// TIA Portal project "liquid refill system" (V18) (continued)
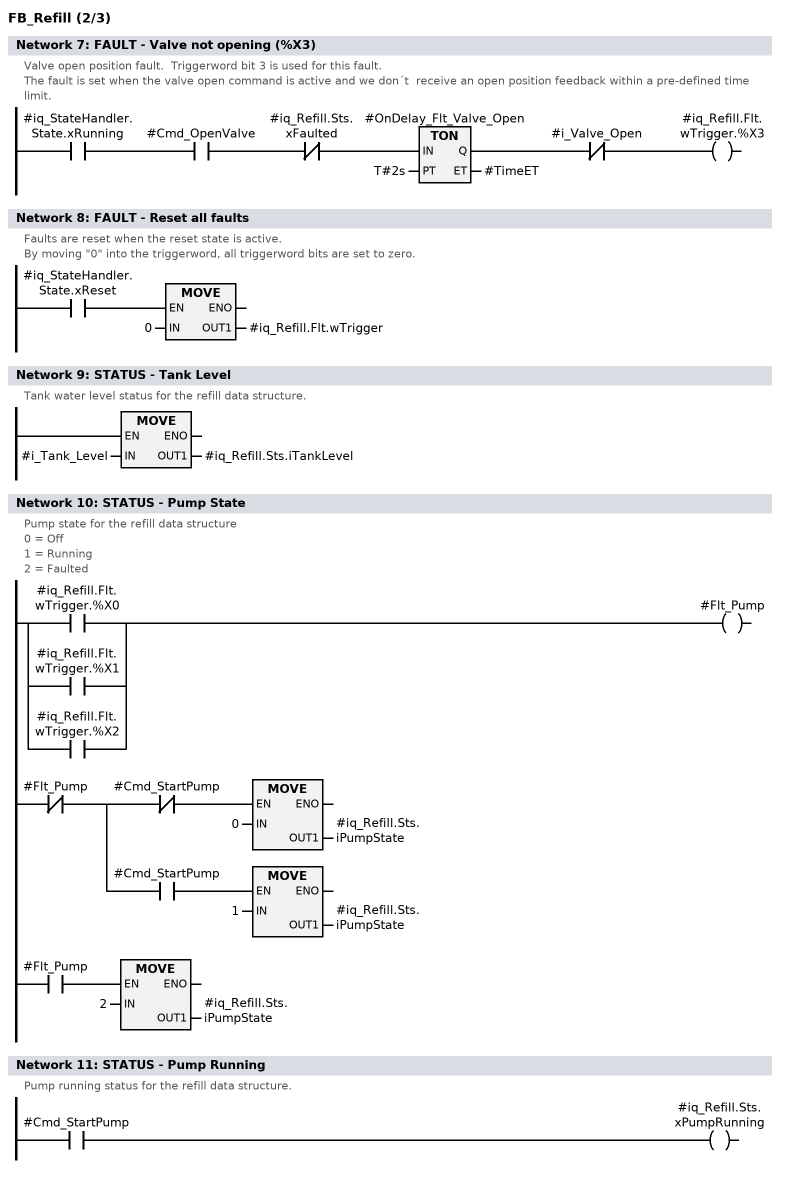
   #OnDelay_Flt_Valve_Open.TON(IN := #iq_StateHandler.State.xRunning AND #Cmd_OpenValve AND NOT #iq_Refill.Sts.xFaulted,
                           PT := T#2s,
                           ET => #TimeET);
   #iq_Refill.Flt.wTrigger.%X3 := #OnDelay_Flt_Valve_Open.Q AND NOT #i_Valve_Open;
END_REGION

REGION Network 8: FAULT - Reset all faults
   // Faults are reset when the reset state is active.
   // By moving "0" into the triggerword, all triggerword bits are set to zero.
   RUNG wire#powerrail
      Contact( #iq_StateHandler.State.xReset )
      Move(in := 0, out1 => #iq_Refill.Flt.wTrigger)
   END_RUNG
   // the same network as SCL:
   IF #iq_StateHandler.State.xReset THEN #iq_Refill.Flt.wTrigger := 0; END_IF;
END_REGION

REGION Network 9: STATUS - Tank Level
   // Tank water level status for the refill data structure.
   RUNG wire#powerrail
      Move(in := #i_Tank_Level, out1 => #iq_Refill.Sts.iTankLevel)
   END_RUNG
   // the same network as SCL:
   #iq_Refill.Sts.iTankLevel := #i_Tank_Level;
END_REGION

REGION Network 10: STATUS - Pump State
   // Pump state for the refill data structure
   // 0 = Off
   // 1 = Running
   // 2 = Faulted
   RUNG wire#powerrail
      Contact( #iq_Refill.Flt.wTrigger.%X0 )
      wire#w1
      Coil( #Flt_Pump )
   END_RUNG
   RUNG wire#powerrail
      Contact( #iq_Refill.Flt.wTrigger.%X1 )
   END_RUNG wire#w1
   RUNG wire#powerrail
      Contact( #iq_Refill.Flt.wTrigger.%X2 )
   END_RUNG wire#w1
   RUNG wire#powerrail
      I_Contact( #Flt_Pump )
      wire#w2
      I_Contact( #Cmd_StartPump )
      Move(in := 0, out1 => #iq_Refill.Sts.iPumpState)
   END_RUNG
   RUNG wire#w2
      Contact( #Cmd_StartPump )
      Move(in := 1, out1 => #iq_Refill.Sts.iPumpState)
   END_RUNG
   RUNG wire#powerrail
      Contact( #Flt_Pump )
      Move(in := 2, out1 => #iq_Refill.Sts.iPumpState)
   END_RUNG
   // the same network as SCL:
   #Flt_Pump := #iq_Refill.Flt.wTrigger.%X0 OR #iq_Refill.Flt.wTrigger.%X1 OR #iq_Refill.Flt.wTrigger.%X2;
   IF NOT #Flt_Pump AND NOT #Cmd_StartPump THEN #iq_Refill.Sts.iPumpState := 0; END_IF;
   IF NOT #Flt_Pump AND #Cmd_StartPump THEN #iq_Refill.Sts.iPumpState := 1; END_IF;
   IF #Flt_Pump THEN #iq_Refill.Sts.iPumpState := 2; END_IF;
END_REGION

REGION Network 11: STATUS - Pump Running
   // Pump running status for the refill data structure.
   RUNG wire#powerrail
      Contact( #Cmd_StartPump )
      Coil( #iq_Refill.Sts.xPumpRunning )
   END_RUNG
   // the same network as SCL:
   #iq_Refill.Sts.xPumpRunning := #Cmd_StartPump;
END_REGION

REGION Network 12: STATUS - Valve State
   // Valve state for the refill data structure
   // 0 = Closed
   // 1 = Open
   // 2 = Faulted
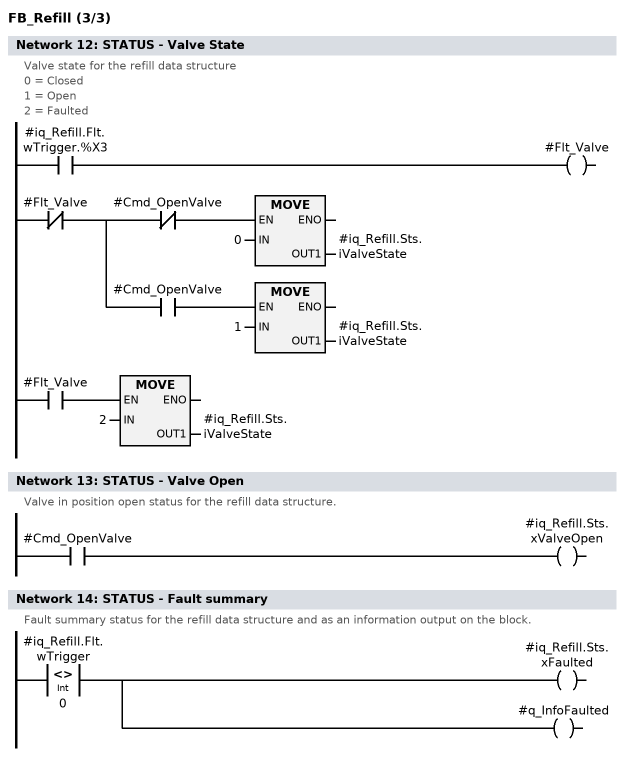
   RUNG wire#powerrail
      Contact( #iq_Refill.Flt.wTrigger.%X3 )
      Coil( #Flt_Valve )
   END_RUNG
   RUNG wire#powerrail
      I_Contact( #Flt_Valve )
      wire#w1
      I_Contact( #Cmd_OpenValve )
      Move(in := 0, out1 => #iq_Refill.Sts.iValveState)
   END_RUNG
   RUNG wire#w1
      Contact( #Cmd_OpenValve )
      Move(in := 1, out1 => #iq_Refill.Sts.iValveState)
   END_RUNG
   RUNG wire#powerrail
      Contact( #Flt_Valve )
      Move(in := 2, out1 => #iq_Refill.Sts.iValveState)
   END_RUNG
   // the same network as SCL:
   #Flt_Valve := #iq_Refill.Flt.wTrigger.%X3;
   IF NOT #Flt_Valve AND NOT #Cmd_OpenValve THEN #iq_Refill.Sts.iValveState := 0; END_IF;
   IF NOT #Flt_Valve AND #Cmd_OpenValve THEN #iq_Refill.Sts.iValveState := 1; END_IF;
   IF #Flt_Valve THEN #iq_Refill.Sts.iValveState := 2; END_IF;
END_REGION

REGION Network 13: STATUS - Valve Open
   // Valve in position open status for the refill data structure.
   RUNG wire#powerrail
      Contact( #Cmd_OpenValve )
      Coil( #iq_Refill.Sts.xValveOpen )
   END_RUNG
   // the same network as SCL:
   #iq_Refill.Sts.xValveOpen := #Cmd_OpenValve;
END_REGION

REGION Network 14: STATUS - Fault summary
   // Fault summary status for the refill data structure and as an information output on the block.
   RUNG wire#powerrail
      { S7_Templates := "SrcType := Int" } NE_Contact(in1 := #iq_Refill.Flt.wTrigger, in2 := 0)
      wire#w1
      Coil( #iq_Refill.Sts.xFaulted )
   END_RUNG
   RUNG wire#w1
      Coil( #q_InfoFaulted )
   END_RUNG
   // the same network as SCL:
   #iq_Refill.Sts.xFaulted := #iq_Refill.Flt.wTrigger <> 0;
   #q_InfoFaulted := #iq_Refill.Sts.xFaulted;
END_REGION
END_FUNCTION_BLOCK

FUNCTION_BLOCK "FB_Supply"   // FB5, LAD
TITLE = EQUIPMENT - Supply
{ S7_Optimized_Access := 'TRUE' }
VERSION : 0.1
// This module consists of a tank with a digital low level sensor, and a valve.
   VAR_INPUT
      i_LevelLow : Bool;
      i_ValveOpen : Bool;
   END_VAR
   VAR_OUTPUT
      q_OpenValve : Bool;
      q_InfoFaulted : Bool;
   END_VAR
   VAR_IN_OUT
      iq_StateHandler : "UDT_Statehandler";
      iq_Supply : "UDT_Supply";
      iq_Refill_Process1 : "UDT_Refill";
      iq_Refill_Process2 : "UDT_Refill";
   END_VAR
   VAR
      OnDelay_LowLvl : IEC_TIMER;
      OnDelay_LowLvlFlt : IEC_TIMER;
      OnDelay_Flt_Valve_Open : IEC_TIMER;
   END_VAR
   VAR_TEMP
      Cmd_OpenValve : Bool;
      TimeTemp : Real;
      TimeET : Time;
      LevelLow : Bool;
      ValveDelayClose : DInt;
      Flt_Valve : Bool;
   END_VAR
BEGIN

REGION Network 1: DELAY - Low Level Signal
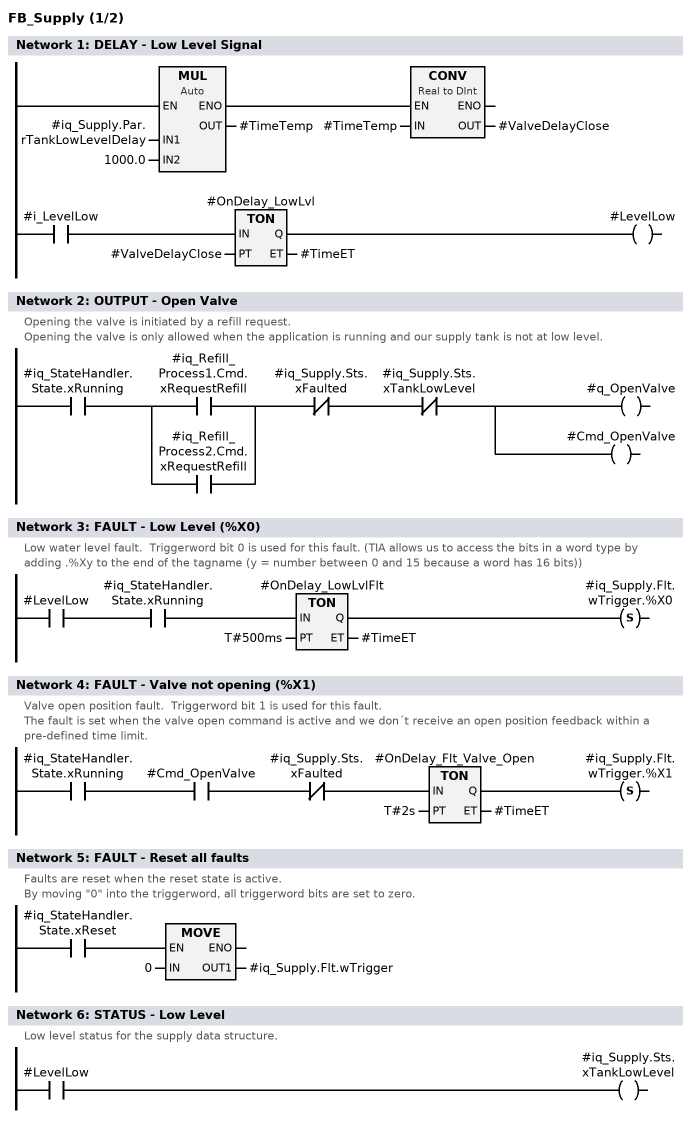
   #TimeTemp := #iq_Supply.Par.rTankLowLevelDelay * 1000.0;
   #ValveDelayClose := REAL_TO_DINT(#TimeTemp);
   #OnDelay_LowLvl.TON(IN := #i_LevelLow, PT := #ValveDelayClose, ET => #TimeET);
   #LevelLow := #OnDelay_LowLvl.Q;
END_REGION

REGION Network 2: OUTPUT - Open Valve
   // Opening the valve is initiated by a refill request.
   // Opening the valve is only allowed when the application is running and our supply tank is not at low level.
   RUNG wire#powerrail
      Contact( #iq_StateHandler.State.xRunning )
      wire#w1
      Contact( #iq_Refill_Process1.Cmd.xRequestRefill )
      wire#w2
      I_Contact( #iq_Supply.Sts.xFaulted )
      I_Contact( #iq_Supply.Sts.xTankLowLevel )
      wire#w3
      Coil( #q_OpenValve )
   END_RUNG
   RUNG wire#w1
      Contact( #iq_Refill_Process2.Cmd.xRequestRefill )
   END_RUNG wire#w2
   RUNG wire#w3
      Coil( #Cmd_OpenValve )
   END_RUNG
   // the same network as SCL:
   #q_OpenValve := #iq_StateHandler.State.xRunning AND (#iq_Refill_Process1.Cmd.xRequestRefill OR #iq_Refill_Process2.Cmd.xRequestRefill) AND NOT #iq_Supply.Sts.xFaulted AND NOT #iq_Supply.Sts.xTankLowLevel;
   #Cmd_OpenValve := #q_OpenValve;
END_REGION

REGION Network 3: FAULT - Low Level (%X0)
   // Low water level fault.  Triggerword bit 0 is used for this fault. (TIA allows us to access the bits in a word type by adding .%Xy to the end of the tagname (y = number between 0 and 15 because a word has 16 bits))
   #OnDelay_LowLvlFlt.TON(IN := #LevelLow AND #iq_StateHandler.State.xRunning, PT := T#500ms, ET => #TimeET);
   IF #OnDelay_LowLvlFlt.Q THEN #iq_Supply.Flt.wTrigger.%X0 := TRUE; END_IF;
END_REGION

REGION Network 4: FAULT - Valve not opening (%X1)
   // Valve open position fault.  Triggerword bit 1 is used for this fault.
   // The fault is set when the valve open command is active and we don´t receive an open position feedback within a pre-defined time limit.
   #OnDelay_Flt_Valve_Open.TON(IN := #iq_StateHandler.State.xRunning AND #Cmd_OpenValve AND NOT #iq_Supply.Sts.xFaulted,
                           PT := T#2s,
                           ET => #TimeET);
   IF #OnDelay_Flt_Valve_Open.Q THEN #iq_Supply.Flt.wTrigger.%X1 := TRUE; END_IF;
END_REGION

REGION Network 5: FAULT - Reset all faults
   // Faults are reset when the reset state is active.
   // By moving "0" into the triggerword, all triggerword bits are set to zero.
   RUNG wire#powerrail
      Contact( #iq_StateHandler.State.xReset )
      Move(in := 0, out1 => #iq_Supply.Flt.wTrigger)
   END_RUNG
   // the same network as SCL:
   IF #iq_StateHandler.State.xReset THEN #iq_Supply.Flt.wTrigger := 0; END_IF;
END_REGION

REGION Network 6: STATUS - Low Level
   // Low level status for the supply data structure.
   RUNG wire#powerrail
      Contact( #LevelLow )
      Coil( #iq_Supply.Sts.xTankLowLevel )
   END_RUNG
   // the same network as SCL:
   #iq_Supply.Sts.xTankLowLevel := #LevelLow;
END_REGION

REGION Network 7: STATUS - Valve State
   // Valve state for the supply data structure
   // 0 = Closed
   // 1 = Open
   // 2 = Faulted
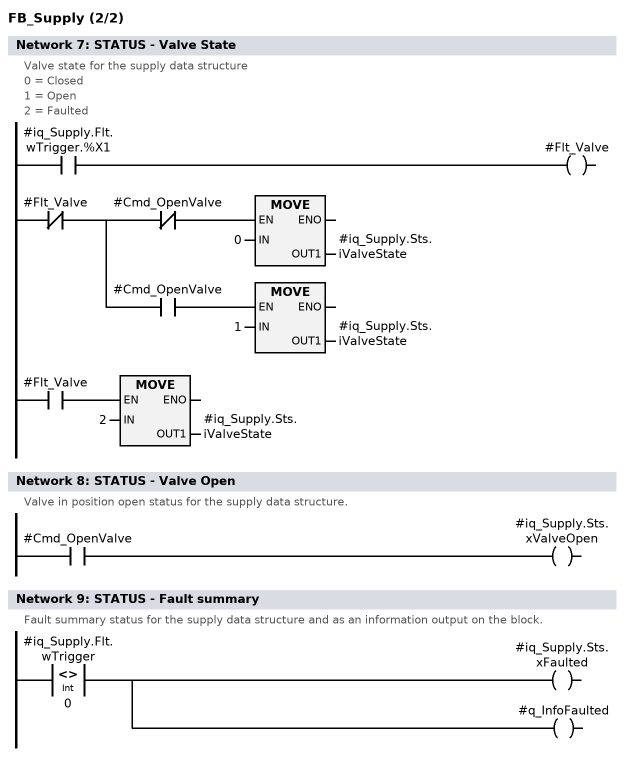
   RUNG wire#powerrail
      Contact( #iq_Supply.Flt.wTrigger.%X1 )
      Coil( #Flt_Valve )
   END_RUNG
   RUNG wire#powerrail
      I_Contact( #Flt_Valve )
      wire#w1
      I_Contact( #Cmd_OpenValve )
      Move(in := 0, out1 => #iq_Supply.Sts.iValveState)
   END_RUNG
   RUNG wire#w1
      Contact( #Cmd_OpenValve )
      Move(in := 1, out1 => #iq_Supply.Sts.iValveState)
   END_RUNG
   RUNG wire#powerrail
      Contact( #Flt_Valve )
      Move(in := 2, out1 => #iq_Supply.Sts.iValveState)
   END_RUNG
   // the same network as SCL:
   #Flt_Valve := #iq_Supply.Flt.wTrigger.%X1;
   IF NOT #Flt_Valve AND NOT #Cmd_OpenValve THEN #iq_Supply.Sts.iValveState := 0; END_IF;
   IF NOT #Flt_Valve AND #Cmd_OpenValve THEN #iq_Supply.Sts.iValveState := 1; END_IF;
   IF #Flt_Valve THEN #iq_Supply.Sts.iValveState := 2; END_IF;
END_REGION

REGION Network 8: STATUS - Valve Open
   // Valve in position open status for the supply data structure.
   RUNG wire#powerrail
      Contact( #Cmd_OpenValve )
      Coil( #iq_Supply.Sts.xValveOpen )
   END_RUNG
   // the same network as SCL:
   #iq_Supply.Sts.xValveOpen := #Cmd_OpenValve;
END_REGION

REGION Network 9: STATUS - Fault summary
   // Fault summary status for the supply data structure and as an information output on the block.
   RUNG wire#powerrail
      { S7_Templates := "SrcType := Int" } NE_Contact(in1 := #iq_Supply.Flt.wTrigger, in2 := 0)
      wire#w1
      Coil( #iq_Supply.Sts.xFaulted )
   END_RUNG
   RUNG wire#w1
      Coil( #q_InfoFaulted )
   END_RUNG
   // the same network as SCL:
   #iq_Supply.Sts.xFaulted := #iq_Supply.Flt.wTrigger <> 0;
   #q_InfoFaulted := #iq_Supply.Sts.xFaulted;
END_REGION
END_FUNCTION_BLOCK

(* ===== HMI "HMI_RT_1" =====
system functions are stored by id; their names below are inferred from use
connection "HMI_Connection_1": ETHERNET, S7_1200_OMS

HMI tags "PLC Machine Tags"
   "Machine_StateHandler" : UDT_Statehandler = PLC "DB - Machine".StateHandler, 1 s

HMI tags "PLC Equipment Tags"
   "Equipment_Supply" : UDT_Supply = PLC "DB - Equipment".Supply, 1 s
   "Equipment_Refill_Process_1" : UDT_Refill = PLC "DB - Equipment".Refill_Process_1 AT %DB1.DBW0, 1 s
   "Equipment_Refill_Process_2" : UDT_Refill = PLC "DB - Equipment".Refill_Process_2 AT %DB1.DBW0, 1 s

HMI tags "Local Template Tags"
   "State_Btn_Overview" : Bool, internal
   "State_Btn_Alarms" : Bool, internal
   "State_Btn_Recipes" : Bool, internal
   "State_Btn_Settings" : Bool, internal
   "iScreenNumber" : Int, internal
   "iRCP_RecordNumber_Actual" : Int, internal
   "sRCP_RecordName_Actual" : WString[254], internal
   "sRCP_RecipeName_Actual" : WString[254], internal
   "Username" : WString[254], internal
   "UserGroupNumber" : Int, internal

HMI tags "PLC Recipe Tags"
   "DB - Equipment_Refill_Process_1_Par_iTankLevelLow(RCP)" : Int = PLC "DB - Equipment".Refill_Process_1.Par.iTankLevelLow, 1 s
   "DB - Equipment_Refill_Process_1_Par_iTankLevelHigh(RCP)" : Int = PLC "DB - Equipment".Refill_Process_1.Par.iTankLevelHigh AT %DB1.DBW0, 1 s
   "DB - Equipment_Refill_Process_2_Par_iTankLevelLow(RCP)" : Int = PLC "DB - Equipment".Refill_Process_2.Par.iTankLevelLow AT %DB1.DBW0, 1 s
   "DB - Equipment_Refill_Process_2_Par_iTankLevelHigh(RCP)" : Int = PLC "DB - Equipment".Refill_Process_2.Par.iTankLevelHigh AT %DB1.DBW0, 1 s
   "DB - Equipment_Supply_Par_rTankLowLevelDelay(RCP)" : Real = PLC "DB - Equipment".Supply.Par.rTankLowLevelDelay AT %DB1.DBW0, 1 s

HMI tags "Local Recipe Tags"
   "iRCP-Number" : Int, internal
   "iRCP-Record Number" : Int, internal

discrete alarms
   1: 'Refill Process1 - Pump - Motor Circuit Breaker Fault', class Errors, trigger "wTrigger" bit 0
   2: 'Refill Process1 - Pump - Local Isolator Fault', class Errors, trigger "wTrigger" bit 1
   3: 'Refill Process1 - Pump - Running Feedback Fault', class Errors, trigger "wTrigger" bit 2
   4: 'Refill Process1 - Valve - Not Opening Fault', class Errors, trigger "wTrigger" bit 3
   5: 'Refill Process2 - Pump - Motor Circuit Breaker Fault', class Errors, trigger "wTrigger" bit 0
   6: 'Refill Process2- Pump - Local Isolator Fault', class Errors, trigger "wTrigger" bit 1
   7: 'Refill Process2 - Pump - Running Feedback Fault', class Errors, trigger "wTrigger" bit 2
   8: 'Refill Process2 - Valve - Not Opening Fault', class Errors, trigger "wTrigger" bit 3
   9: 'Supply- Tank - Low Level Fault', class Errors, trigger "wTrigger" bit 4
   10: 'Supply - Valve - Not Opening Fault', class Errors, trigger "wTrigger" bit 5

text list "Text_ScreenNames": 1 'Process Overview'; 5 'Alarms'; 10 'Recipes'; 20 'Settings'; 6 'Alarm Buffer'; 7 'Diagnostcis'

graphic list "GraphicList_Btn_Template_Overview": 0 'Btn_Template_Overview_Off'; 1 'Btn_Template_Overview_On'

graphic list "GraphicList_Btn_Template_Alarms": 0 'Btn_Template_Alarm_Off'; 1 'Btn_Template_Alarm_On'

graphic list "GraphicList_Btn_Template_Recipes": 0 'Btn_Template_Rcp_Off'; 1 'Btn_Template_Rcp_On'

graphic list "GraphicList_Btn_Template_Settings": 0 'Btn_Template_Settings_Off'; 1 'Btn_Template_Settings_On'

graphic list "GraphicList_Pump_State": 0 'Process_Pump_Off'; 1 'Process_Pump_On'; 2 'Process_Pump_Flt'

graphic list "GraphicList_Valve_State": 0 'Process_Valve_Off'; 1 'Process_Valve_On'; 2 'Process_Valve_Flt'

recipe "Recipe-Equipment": Refill Process 1 - Tank Level High <- "DB - Equipment_Refill_Process_1_Par_iTankLevelHigh(RCP)", Refill Process 2 - Tank Level High <- "DB - Equipment_Refill_Process_2_Par_iTankLevelHigh(RCP)", Supply - Low level Delay <- "DB - Equipment_Supply_Par_rTankLowLevelDelay(RCP)", Refill Process 1 - Tank Level low <- "DB - Equipment_Refill_Process_1_Par_iTankLevelLow(RCP)", Refill Process 2 - Tank Level low <- "DB - Equipment_Refill_Process_2_Par_iTankLevelLow(RCP)"

Template "Template_1" 800x480
   GraphicView "Template_Graphic view_1" at 0,0 size 800x480; Picture "Background_Template"
   Rectangle "Template_Rectangle_1" at 0,0 size 108x38
      Appearance <- "UserGroupNumber"
   Rectangle "Template_Rectangle_4" at 3,43 size 689x434
      Appearance <- "iState"
   Button "Template_Button_1" at 696,1 size 104x78; TextOff 'Text'; PictureList "GraphicList_Btn_Template_Overview"
      ProcessValue <- "State_Btn_Overview"
      on Release: ActivateScreen("1 Overview", 0)
   Button "Template_Button_2" at 696,75 size 104x78; TextOff 'Text'; PictureList "GraphicList_Btn_Template_Alarms"
      on Release: ActivateScreen("5 Alarms", 0)
      ProcessValue <- "State_Btn_Alarms"
   Button "Template_Button_3" at 696,150 size 104x78; TextOff 'Text'; PictureList "GraphicList_Btn_Template_Recipes"
      on Release: ActivateScreen("10 Recipes", 0)
      ProcessValue <- "State_Btn_Recipes"
   Button "Template_Button_4" at 696,223 size 104x78; TextOff 'Text'; PictureList "GraphicList_Btn_Template_Settings"
      on Release: ActivateScreen("20 Settings", 0)
      ProcessValue <- "State_Btn_Settings"
   Button "Template_Button_5" at 696,305 size 104x85; TextOff 'Text'; PictureList "GraphicList_Btn_Template_Overview"; PictureOff "Btn_Template_Start_Off"; PictureOn "Btn_Template_Start_On"; Authorization "Operation"
      ProcessValue <- "State_Btn_Overview"
      on Press: function_b14e0dd5("xStart", 0)
   Button "Template_Button_6" at 696,397 size 104x78; TextOff 'Text'; PictureList "GraphicList_Btn_Template_Overview"; PictureOff "Btn_Template_Stop_Off"; PictureOn "Btn_Template_Stop_On"; Authorization "Operation"
      on Press: function_b14e0dd5("xStop", 0)
      ProcessValue <- "State_Btn_Overview"
   SymbolicIOField "Template_Symbolic I/O field_1" at 111,0 size 234x38; TextOff '0'; TextOn '1'; TextList "Text_ScreenNames"
      ProcessValue <- "iScreenNumber"
   DateTimeField "Template_Date/time field_1" at 480,0 size 219x38
   TextField "Template_Text field_2" at 375,7 size 14x26; Text '-'
   IOField "Template_I/O field_1" at 347,7 size 29x22; FormatPattern 99
      ProcessValue <- "iRCP_RecordNumber_Actual"
   IOField "Template_I/O field_2" at 363,7 size 135x22; FormatPattern ????????
      ProcessValue <- "sRCP_RecordName_Actual"
   IOField "Template_I/O field_3" at 0,0 size 111x40; FormatPattern ????????
      ProcessValue <- "Username"

screen "1 Overview" 800x480, template "Template_1"
   on GenerateScreen: SetBit("State_Btn_Overview"); SetTag("iScreenNumber", 1)
   on ClearScreen: ResetBit("State_Btn_Overview")
   GraphicView "Graphic view_1" at 31,306 size 137x147; Picture "Process_Tank_Supply"
   GraphicView "Graphic view_2" at 471,110 size 137x147; Picture "Process_Tank_Refill"
   GraphicView "Graphic view_3" at 473,303 size 137x147; Picture "Process_Tank_Refill"
   Line "Line_2" at 99,184 size 162x0
      Appearance <- "xValveOpen"
   Line "Line_3" at 263,180 size 0x99
      Appearance <- "xValveOpen"
   Line "Line_5" at 263,281 size 239x0
      Appearance <- "xValveOpen"
   Line "Line_4" at 264,91 size 239x0
      Appearance <- "xValveOpen"
   Line "Line_6" at 504,91 size 0x19
      Appearance <- "xValveOpen"
   Line "Line_7" at 502,282 size 0x20
      Appearance <- "xValveOpen"
   Line "Line_8" at 263,91 size 0x89
      Appearance <- "xValveOpen"
   TextField "Text field_1" at 113,283 size 93x20; Text 'Supply Tank'
   TextField "Text field_2" at 511,84 size 116x20; Text 'Process Tank 1'
   TextField "Text field_3" at 511,278 size 116x20; Text 'Process Tank 2'
   TextField "Text field_4" at 283,113 size 58x20; Text 'Pump 1'
   TextField "Text field_5" at 276,304 size 58x20; Text 'Pump 2'
   TextField "Text field_6" at 371,111 size 60x20; Text 'Valve 1'
   TextField "Text field_7" at 374,303 size 60x20; Text 'Valve 2'
   TextField "Text field_8" at 155,200 size 51x20; Text 'Valve'
   GraphicIOField "Graphic I/O field_1" at 287,71 size 38x40; PictureList "GraphicList_Pump_State"
      ProcessValue <- "iPumpState"
   GraphicIOField "Graphic I/O field_2" at 287,262 size 38x40; PictureList "GraphicList_Pump_State"
      ProcessValue <- "iPumpState"
   GraphicIOField "Graphic I/O field_3" at 376,66 size 53x39; PictureList "GraphicList_Valve_State"
      ProcessValue <- "iValveState"
   GraphicIOField "Graphic I/O field_4" at 376,256 size 53x39; PictureList "GraphicList_Valve_State"
      ProcessValue <- "iValveState"
   GraphicIOField "Graphic I/O field_5" at 156,160 size 53x39; PictureList "GraphicList_Valve_State"
      ProcessValue <- "iValveState"
   Bar "Bar_1" at 482,111 size 115x106; MinimumValue 0; MaximumValue 100
      ProcessValue <- "iTankLevel"
   Bar "Bar_2" at 484,302 size 115x106; MinimumValue 0; MaximumValue 100
      ProcessValue <- "iTankLevel"
   Rectangle "Rectangle_1" at 42,328 size 115x84
      Visibility <- "xTankLowLevel"
   Line "Line_9" at 35,416 size 131x1
      Appearance <- "xValveOpen"
   IOField "I/O field_1" at 606,217 size 59x32; Authorization "Operation"; FormatPattern 999; Unit %
      ProcessValue <- "iTankLevelLow"
   TextField "Text field_9" at 617,189 size 36x22; Text 'Low'
   Group "Low1" at 606,189 size 59x60; Authorization "Operation"
   Group "High1" at 606,107 size 59x60; Authorization "Operation"
   Group "High2" at 608,299 size 59x60; Authorization "Operation"
   Group "Low2" at 608,381 size 59x60; Authorization "Operation"
   Group "Low2_1" at 169,376 size 59x60; Authorization "Operation"; FormatPattern 999; Unit %
   IOField "I/O field_3" at 606,135 size 59x32; Authorization "Operation"; FormatPattern 999; Unit %
      ProcessValue <- "iTankLevelHigh"
   TextField "Text field_11" at 617,107 size 39x22; Text 'High'
   IOField "I/O field_4" at 608,327 size 59x32; Authorization "Operation"; FormatPattern 999; Unit %
      ProcessValue <- "iTankLevelHigh"
   TextField "Text field_12" at 619,299 size 39x22; Text 'High'
   IOField "I/O field_2" at 608,409 size 59x32; Authorization "Operation"; FormatPattern 999; Unit %
      ProcessValue <- "iTankLevelLow"
   TextField "Text field_10" at 619,381 size 36x22; Text 'Low'
   IOField "I/O field_5" at 169,404 size 59x32; Authorization "Operation"; FormatPattern 99.9; Unit s
      ProcessValue <- "rTankLowLevelDelay"
   TextField "Text field_13" at 180,376 size 36x22; Text 'Low'

screen "5 Alarms" 800x480, template "Template_1"
   on GenerateScreen: SetBit("State_Btn_Alarms"); SetTag("iScreenNumber", 5)
   on ClearScreen: ResetBit("State_Btn_Alarms")
   AlarmView "Alarm view_1" at 7,48 size 604x423
   Button "Template_Button_6" at 613,397 size 71x72; TextOff 'Text'; PictureList "GraphicList_Btn_Template_Overview"; PictureOff "Btn_Reset_Off"; PictureOn "Btn_Reset_On"; Authorization "Operation"
      on Press: function_b14e0dd5("xReset", 0)
      ProcessValue <- "State_Btn_Overview"
   Button "Template_Button_1" at 613,50 size 72x72; TextOff 'Text'; PictureList "GraphicList_Btn_Template_Overview"; PictureOff "Btn_AlarmBuffer_Off"; PictureOn "Btn_AlarmBuffer_On"
      ProcessValue <- "State_Btn_Overview"
      on Release: ActivateScreen("6 Alarm Buffer", 0)
   Button "Template_Button_2" at 614,126 size 72x72; TextOff 'Text'; PictureList "GraphicList_Btn_Template_Overview"; PictureOff "Btn_Diagnostics_Off"; PictureOn "Btn_Diagnostics_On"
      on Release: ActivateScreen("7 Diagnostics", 0)
      ProcessValue <- "State_Btn_Overview"

screen "10 Recipes" 800x480, template "Template_1"
   on GenerateScreen: SetBit("State_Btn_Recipes"); SetTag("iScreenNumber", 10)
   on ClearScreen: ResetBit("State_Btn_Recipes")
   RecipeView "Recipe view_1" at 9,50 size 600x419; Recipe "Recipe-Equipment"; Tag4RecipeNumber "iRCP-Number"; Tag4DataRecord "iRCP-Record Number"; Authorization "Supervision"
   Button "Template_Button_1" at 613,50 size 72x72; TextOff 'Text'; PictureList "GraphicList_Btn_Template_Overview"; PictureOff "Btn_Load_Rcp_Off"; PictureOn "Btn_Load_Rcp_On"; Authorization "Supervision"
      ProcessValue <- "State_Btn_Overview"
      on Press: function_bbf3fe93("Recipe-Equipment", N)
      on Release: SetTag("iRCP_RecordNumber_Actual", "iRCP-Record Number"); function_b69f32de("Recipe-Equipment", "iRCP-Record Number", "sRCP_RecipeName_Actual", "sRCP_RecordName_Actual", N)

screen "20 Settings" 800x480, template "Template_1"
   on GenerateScreen: SetBit("State_Btn_Settings"); SetTag("iScreenNumber", 20)
   on ClearScreen: ResetBit("State_Btn_Settings")
   Button "Template_Button_1" at 47,127 size 72x72; TextOff 'Text'; PictureList "GraphicList_Btn_Template_Overview"; PictureOff "Btn_Calibrate_Off"; PictureOn "Btn_Calibrate_On"; Authorization "Maintenance"
      ProcessValue <- "State_Btn_Overview"
      on Release: function_bc3e350c()
   TextField "Text field_1" at 48,199 size 72x20; Text 'Calibrate'
   Button "Template_Button_2" at 182,128 size 72x72; TextOff 'Text'; PictureList "GraphicList_Btn_Template_Overview"; PictureOff "Btn_CleanScreen_Off"; PictureOn "Btn_CleanScreen_On"; Authorization "Operation"
      on Release: function_bc3e350c()
      ProcessValue <- "State_Btn_Overview"
      on Click: function_be740847(15)
   TextField "Text field_2" at 195,200 size 45x20; Text 'Clean'
   Button "Template_Button_3" at 49,238 size 72x72; TextOff 'Text'; PictureList "GraphicList_Btn_Template_Overview"; PictureOn "Btn_LogOff_On"; PictureOff "Btn_LogOff_Off"
      on Release: function_bc3e350c()
      ProcessValue <- "State_Btn_Overview"
      on Click: function_f23ef4c9()
   TextField "Text field_3" at 54,310 size 58x20; Text 'Log Off'
   Group "Group_2" at 49,238 size 72x92; PictureList "GraphicList_Btn_Template_Overview"; PictureOff "Btn_Calibrate_Off"; PictureOn "Btn_Calibrate_On"
   Group "Group_3" at 182,238 size 72x92; PictureList "GraphicList_Btn_Template_Overview"; PictureOff "Btn_Calibrate_Off"; PictureOn "Btn_Calibrate_On"; Authorization "Maintenance"
   Group "Group_1" at 182,128 size 72x92; PictureList "GraphicList_Btn_Template_Overview"; PictureOff "Btn_Calibrate_Off"; PictureOn "Btn_Calibrate_On"; Authorization "Operation"
   Group "Group" at 47,127 size 73x92; PictureList "GraphicList_Btn_Template_Overview"; PictureOff "Btn_Calibrate_Off"; PictureOn "Btn_Calibrate_On"; Authorization "Maintenance"
   TextField "Text field_5" at 310,118 size 114x20; Text 'Project Name :'
   TextField "Text field_6" at 310,146 size 99x20; Text 'Created On :'
   TextField "Text field_7" at 310,172 size 68x20; Text 'Author :'
   TextField "Text field_8" at 310,199 size 100x20; Text 'Description :'
   TextField "Text field_9" at 446,118 size 61x20; Text 'Refill'
   TextField "Text field_10" at 446,146 size 128x20; Text 'January 27 2026'
   TextField "Text field_11" at 446,173 size 106x20; Text 'Sobhan Sahaf'
   TextField "Text field_12" at 452,208 size 331x90; Text 'This refill application consists of 1 supply tank and 2 process tanks. a process tank can be refilled with liquid from the supply tank using the appropriate pump and valves .'
   TextField "Text field_13" at 310,356 size 136x20; Text 'PLC Device Type :'
   TextField "Text field_14" at 310,382 size 138x20; Text 'HMI Device Type :'
   TextField "Text field_15" at 310,409 size 138x20; Text 'Connection Type :'
   TextField "Text field_16" at 446,356 size 124x20; Text 'Simatic S7-1200'
   TextField "Text field_17" at 446,384 size 112x20; Text 'TP900 Comfort'
   TextField "Text field_18" at 446,411 size 65x20; Text 'Profinet'
   Button "Template_Button_4" at 182,238 size 72x72; TextOff 'Text'; PictureList "GraphicList_Btn_Template_Overview"; PictureOff "Btn_StopRuntime_Off"; PictureOn "Btn_StopRuntime_On"; Authorization "Maintenance"
      on Release: function_bc3e350c()
      ProcessValue <- "State_Btn_Overview"
      on Click: StopRuntime(0)
   TextField "Text field_4" at 202,310 size 32x20; Text 'Exit'
   TextField "Text field_19" at 306,84 size 151x20; Text 'Project Information'
   TextField "Text field_20" at 306,324 size 151x20; Text 'System Information'
   TextField "Text field_21" at 21,84 size 108x20; Text 'HMI Functions'

screen "6 Alarm Buffer" 800x480, template "Template_1"
   on GenerateScreen: SetBit("State_Btn_Alarms"); SetTag("iScreenNumber", 6)
   on ClearScreen: ResetBit("State_Btn_Alarms")
   AlarmView "Alarm view_1" at 7,48 size 604x423
   Button "Template_Button_6" at 613,51 size 72x72; TextOff 'Text'; PictureList "GraphicList_Btn_Template_Overview"; PictureOff "Btn_PreviousScreen_Off"; PictureOn "Btn_PreviousScreen_On"
      ProcessValue <- "State_Btn_Overview"
      on Release: function_efd93a16()

screen "7 Diagnostics" 800x480, template "Template_1"
   on GenerateScreen: SetBit("State_Btn_Alarms"); SetTag("iScreenNumber", 7)
   on ClearScreen: ResetBit("State_Btn_Alarms")
   Button "Template_Button_6" at 613,51 size 72x72; TextOff 'Text'; PictureList "GraphicList_Btn_Template_Overview"; PictureOff "Btn_PreviousScreen_Off"; PictureOn "Btn_PreviousScreen_On"
      on Release: function_efd93a16()
      ProcessValue <- "State_Btn_Overview"
   SysDiagControl "System diagnostics view_1" at 8,49 size 600x421

scheduled task "UserName"
   on Action: function_f41c6f6c("Username"); function_e1ab61de("UserGroupNumber")
*)